   
   //M214
   M2xx_CONVEYOR[11].INPUT_xProtectionRot := A152AP1:3:I.Pt08.Data;
   M2xx_CONVEYOR[11].INPUT_xProtectionFan := xAlwaysON;
   M2xx_CONVEYOR[11].INPUT_xLocalSafetySwitch := A152AP1:10:I.Pt00.Data;
   M2xx_CONVEYOR[11].INPUT_xThermalProbe := A152AP1:10:I.Pt01.Data;
   M2xx_CONVEYOR[11].INPUT_xDriveInhibit := M214_M1_DR.CIPAxisState = 9;
   M2xx_CONVEYOR[11].INPUT_xDriveReady := M214_M1_DR.ServoActionStatus;
   M2xx_CONVEYOR[11].INPUT_xDriveError := M214_M1_DR.AxisFault <> 0 OR M214_M1_DR.ModuleFaults <> 0;
   M2xx_CONVEYOR[11].INPUT_xRotationFeedback := M214_M1_DR.MotionStatus <> 0;
   
   //M215
   M2xx_CONVEYOR[12].INPUT_xProtectionRot := A152AP1:3:I.Pt09.Data;
   M2xx_CONVEYOR[12].INPUT_xProtectionFan := xAlwaysON;
   M2xx_CONVEYOR[12].INPUT_xLocalSafetySwitch := A152AP1:10:I.Pt02.Data;
   M2xx_CONVEYOR[12].INPUT_xThermalProbe := A152AP1:10:I.Pt03.Data;
   M2xx_CONVEYOR[12].INPUT_xDriveInhibit := M215_M1_DR.CIPAxisState = 9;
   M2xx_CONVEYOR[12].INPUT_xDriveReady := M215_M1_DR.ServoActionStatus;
   M2xx_CONVEYOR[12].INPUT_xDriveError := M215_M1_DR.AxisFault <> 0 OR M215_M1_DR.ModuleFaults <> 0;
   M2xx_CONVEYOR[12].INPUT_xRotationFeedback := M215_M1_DR.MotionStatus <> 0;
   
   //M216
   M2xx_CONVEYOR[13].INPUT_xProtectionRot := A152AP1:3:I.Pt10.Data;
   M2xx_CONVEYOR[13].INPUT_xProtectionFan := xAlwaysON;
   M2xx_CONVEYOR[13].INPUT_xLocalSafetySwitch := A152AP1:10:I.Pt04.Data;
   M2xx_CONVEYOR[13].INPUT_xThermalProbe := A152AP1:10:I.Pt05.Data;
   M2xx_CONVEYOR[13].INPUT_xDriveInhibit := M216_M1_DR.CIPAxisState = 9;
   M2xx_CONVEYOR[13].INPUT_xDriveReady := M216_M1_DR.ServoActionStatus;
   M2xx_CONVEYOR[13].INPUT_xDriveError := M216_M1_DR.AxisFault <> 0 OR M216_M1_DR.ModuleFaults <> 0;
   M2xx_CONVEYOR[13].INPUT_xRotationFeedback := M216_M1_DR.MotionStatus <> 0;
   
   //M217
   M2xx_CONVEYOR[14].INPUT_xProtectionRot := A152AP1:3:I.Pt11.Data;
   M2xx_CONVEYOR[14].INPUT_xProtectionFan := xAlwaysON;
   M2xx_CONVEYOR[14].INPUT_xLocalSafetySwitch := A152AP1:10:I.Pt06.Data;
   M2xx_CONVEYOR[14].INPUT_xThermalProbe := A152AP1:10:I.Pt07.Data;
   M2xx_CONVEYOR[14].INPUT_xDriveInhibit := M217_M1_DR.CIPAxisState = 9;
   M2xx_CONVEYOR[14].INPUT_xDriveReady := M217_M1_DR.ServoActionStatus;
   M2xx_CONVEYOR[14].INPUT_xDriveError := M217_M1_DR.AxisFault <> 0 OR M217_M1_DR.ModuleFaults <> 0;
   M2xx_CONVEYOR[14].INPUT_xRotationFeedback := M217_M1_DR.MotionStatus <> 0;
   
   //M218
   M2xx_CONVEYOR[15].INPUT_xProtectionRot := A152AP1:3:I.Pt12.Data;
   M2xx_CONVEYOR[15].INPUT_xProtectionFan := xAlwaysON;
   M2xx_CONVEYOR[15].INPUT_xLocalSafetySwitch := A152AP1:10:I.Pt08.Data;
   M2xx_CONVEYOR[15].INPUT_xThermalProbe := A152AP1:10:I.Pt09.Data;
   M2xx_CONVEYOR[15].INPUT_xDriveInhibit := M218_M1_DR.CIPAxisState = 9;
   M2xx_CONVEYOR[15].INPUT_xDriveReady := M218_M1_DR.ServoActionStatus;
   M2xx_CONVEYOR[15].INPUT_xDriveError := M218_M1_DR.AxisFault <> 0 OR M218_M1_DR.ModuleFaults <> 0;
   M2xx_CONVEYOR[15].INPUT_xRotationFeedback := M218_M1_DR.MotionStatus <> 0;
   
   //M219
   M2xx_CONVEYOR[16].INPUT_xProtectionRot := A152AP1:3:I.Pt13.Data;
   M2xx_CONVEYOR[16].INPUT_xProtectionFan := xAlwaysON;
   M2xx_CONVEYOR[16].INPUT_xLocalSafetySwitch := A152AP1:10:I.Pt10.Data;
   M2xx_CONVEYOR[16].INPUT_xThermalProbe := A152AP1:10:I.Pt11.Data;
   M2xx_CONVEYOR[16].INPUT_xDriveInhibit := M219_M1_DR.CIPAxisState = 9;
   M2xx_CONVEYOR[16].INPUT_xDriveReady := M219_M1_DR.ServoActionStatus;
   M2xx_CONVEYOR[16].INPUT_xDriveError := M219_M1_DR.AxisFault <> 0 OR M219_M1_DR.ModuleFaults <> 0;
   M2xx_CONVEYOR[16].INPUT_xRotationFeedback := M219_M1_DR.MotionStatus <> 0;
   
   //M301M1
   M2xx_CONVEYOR[17].INPUT_xProtectionRot := A152AP1:3:I.Pt14.Data;
   M2xx_CONVEYOR[17].INPUT_xProtectionFan := xAlwaysON;
   M2xx_CONVEYOR[17].INPUT_xLocalSafetySwitch := A152AP1:10:I.Pt12.Data;
   M2xx_CONVEYOR[17].INPUT_xThermalProbe := A152AP1:10:I.Pt13.Data;
   M2xx_CONVEYOR[17].INPUT_xDriveInhibit := M301_M1_DR.CIPAxisState = 9;
   M2xx_CONVEYOR[17].INPUT_xDriveReady := M301_M1_DR.ServoActionStatus;
   M2xx_CONVEYOR[17].INPUT_xDriveError := M301_M1_DR.AxisFault <> 0 OR M301_M1_DR.ModuleFaults <> 0;
   M2xx_CONVEYOR[17].INPUT_xRotationFeedback := M301_M1_DR.MotionStatus <> 0;
   
   
   //M301M2
   M2xx_CONVEYOR[18].INPUT_xProtectionRot := A152AP1:3:I.Pt15.Data;
   M2xx_CONVEYOR[18].INPUT_xProtectionFan := xAlwaysON;
   M2xx_CONVEYOR[18].INPUT_xLocalSafetySwitch := A152AP1:10:I.Pt14.Data;
   M2xx_CONVEYOR[18].INPUT_xThermalProbe := A152AP1:10:I.Pt15.Data;
   M2xx_CONVEYOR[18].INPUT_xDriveInhibit := M301_M2_DR.CIPAxisState = 9;
   M2xx_CONVEYOR[18].INPUT_xDriveReady := M301_M2_DR.ServoActionStatus;
   M2xx_CONVEYOR[18].INPUT_xDriveError := M301_M2_DR.AxisFault <> 0 OR M301_M2_DR.ModuleFaults <> 0;
   M2xx_CONVEYOR[18].INPUT_xRotationFeedback := M301_M2_DR.MotionStatus <> 0;
   
   
   //M220
   M2xx_CONVEYOR[19].INPUT_xProtectionRot := A152AP1:4:I.Pt00.Data;
   M2xx_CONVEYOR[19].INPUT_xProtectionFan := xAlwaysON;
   M2xx_CONVEYOR[19].INPUT_xLocalSafetySwitch := A152AP1:11:I.Pt00.Data;
   M2xx_CONVEYOR[19].INPUT_xThermalProbe := A152AP1:11:I.Pt01.Data;
   M2xx_CONVEYOR[19].INPUT_xDriveInhibit := M220_M1_DR.CIPAxisState = 9;
   M2xx_CONVEYOR[19].INPUT_xDriveReady := M220_M1_DR.ServoActionStatus;
   M2xx_CONVEYOR[19].INPUT_xDriveError := M220_M1_DR.AxisFault <> 0 OR M220_M1_DR.ModuleFaults <> 0;
   M2xx_CONVEYOR[19].INPUT_xRotationFeedback := M220_M1_DR.MotionStatus <> 0;
   
   
   // MAPPING PREVIOUS PROGRAM INPUTS
   
   //ALARM RESET
   I[16].9 := A152AP1:11:I.Pt08.Data;; //VMCC MB Alarm Silence
   I[16].10 := A152AP1:11:I.Pt09.Data;; //VMCC MB Alarm Reset
   
   //ISRA 5D
   I[16].0 := A152AP1:12:I.Pt00.Data; //ISRA 5D 24 VDC OK
   I[16].4 := A152AP1:11:I.Pt06.Data; //ISRA 5D 12 VDC OK
   I[16].5 := A152AP1:11:I.Pt07.Data; //ISRA 5D SYSTEM OK
   I[16].6 := A152AP1:11:I.Pt15.Data; //ISRA 5D System Warning
   I[16].7 := A152AP1:11:I.Pt12.Data; //ISRA 5D System Error 1
   I[16].8 := A152AP1:11:I.Pt13.Data; //ISRA 5D System Error 2
   I[16].14 := A152AP1:11:I.Pt14.Data; //ISRA 5D System Crossbreak
   
   //CHILLED WATER & SUB SURFACE
   I[17].1 := A152AP1:12:I.Pt01.Data; //South Chilled Water Blower Off PB I02105
   I[17].2 := A152AP1:12:I.Pt02.Data; //North Subsurface Cutter Alarm Signal
   I[17].3 := A152AP1:12:I.Pt03.Data; //South Subsurface Cutter Alarm Signal
   I[17].4 := A152AP1:12:I.Pt04.Data; //South Chilled Water Blower On PB I02104
   I[17].5 := A152AP1:12:I.Pt05.Data; //South Chilled Water Blower Off PB I02105
   I[17].7 := A152AP1:12:I.Pt07.Data; //South Chilled Water Blower VFD is Running Without Faults
   I[17].10 := A152AP1:12:I.Pt10.Data; //North Chilled Water Blower On PB I02112
   I[17].11 := A152AP1:12:I.Pt11.Data; //North Chilled Water Blower Off PB I02113
   I[17].13 := A152AP1:12:I.Pt13.Data; //North Chilled Water Blower VFD is Running Without Faults
   
   // CROSSBREAK ZONE 1
   I[24].0 := CB_1CS:0:I.0; //CRSSBRK ZONE 1 North Outside Bypass Switch
   I[24].1 := CB_1CS:0:I.1; //CRSSBRK ZONE 1 North Inside Bypass Switch
   I[24].2 := CB_1CS:0:I.2; //CRSSBRK ZONE 1 South Outside Bypass Switch
   I[24].3 := CB_1CS:0:I.3; //CRSSBRK ZONE 1 South Inside Bypass Switch
   I[24].4 := CB_1CS:0:I.4; //CRSSBRK ZONE 1 North Outside Photo-cell
   I[24].5 := CB_1CS:0:I.5; //CRSSBRK ZONE 1 North Inside Photo-cell
   I[24].6 := CB_1CS:0:I.6; //CRSSBRK ZONE 1 South Outside Photo-cell
   I[24].7 := CB_1CS:0:I.7; //CRSSBRK ZONE 1 South Inside Photo-cell
   I[24].8 := CB_1CS:0:I.8; //Cullet System M37B Fwd Direction Selector (Outside)
   I[24].9 := CB_1CS:0:I.9; //Cullet System M37B Rev Direction Selector (Outside)
   I[24].10 := CB_1CS:0:I.10; //Cullet System M47B Fwd Direction Selector (Outside)
   I[24].11 := CB_1CS:0:I.11; //Cullet System M47B Rev Direction Selector (Outside)
   I[24].12 := CB_1CS:0:I.12; //Diverter Position Selector At Cullet Op Panel (Input from cullet belts 51 running)
   I[24].13 := CB_1CS:0:I.13; //(Input from cullet belts 52 running)
   I[24].14 := CB_1CS:0:I.14; //spare
   I[24].15 := CB_1CS:0:I.15; //spare
   
   // CROSSBREAK ZONE 2
   I[26].0 := CB_2CS:0:I.0; //CRSSBRK ZONE 2 North Outside Bypass Switch
   I[26].1 := CB_2CS:0:I.1; //CRSSBRK ZONE 2 North Inside Bypass Switch
   I[26].2 := CB_2CS:0:I.2; //CRSSBRK ZONE 2 South Outside Bypass Switch
   I[26].3 := CB_2CS:0:I.3; //CRSSBRK ZONE 2 South Inside Bypass Switch
   I[26].4 := CB_2CS:0:I.4; //CRSSBRK ZONE 2 North Outside Photo-cell
   I[26].5 := CB_2CS:0:I.5; //CRSSBRK ZONE 2 North Inside Photo-cell
   I[26].6 := CB_2CS:0:I.6; //CRSSBRK ZONE 2 South Outside Photo-cell
   I[26].7 := CB_2CS:0:I.7; //CRSSBRK ZONE 2 South Inside Photo-cell
   I[26].8 := CB_2CS:0:I.8; //spare
   I[26].9 := CB_2CS:0:I.9; //spare
   I[26].10 := CB_2CS:0:I.10; //spare
   I[26].11 := CB_2CS:0:I.11; //spare
   I[26].12 := CB_2CS:0:I.12; //spare
   I[26].13 := CB_2CS:0:I.13; //Adapter power ON
   I[26].14 := CB_2CS:0:I.14; //Input power ON
   I[26].15 := CB_2CS:0:I.15; //Output power ON
   
   // CROSSBREAK ZONE 3
   I[28].0 := CB_3CS:0:I.0; //CRSSBRK ZONE 3 North Outside Bypass Switch
   I[28].1 := CB_3CS:0:I.1; //CRSSBRK ZONE 3 North Inside Bypass Switch
   I[28].2 := CB_3CS:0:I.2; //CRSSBRK ZONE 3 South Outside Bypass Switch
   I[28].3 := CB_3CS:0:I.3; //CRSSBRK ZONE 3 South Inside Bypass Switch
   I[28].4 := CB_3CS:0:I.4; //CRSSBRK ZONE 3 North Outside Photo-cell
   I[28].5 := CB_3CS:0:I.5; //CRSSBRK ZONE 3 North Inside Photo-cell
   I[28].6 := CB_3CS:0:I.6; //CRSSBRK ZONE 3 South Outside Photo-cell
   I[28].7 := CB_3CS:0:I.7; //CRSSBRK ZONE 3 South Inside Photo-cell
   I[28].8 := CB_3CS:0:I.8; //spare
   I[28].9 := CB_3CS:0:I.9; //spare
   I[28].10 := CB_3CS:0:I.10; //spare
   I[28].11 := CB_3CS:0:I.11; //spare
   I[28].12 := CB_3CS:0:I.12; //spare
   I[28].13 := CB_3CS:0:I.13; //Adapter power ON
   I[28].14 := CB_3CS:0:I.14; //Input power ON
   I[28].15 := CB_3CS:0:I.15; //Output power ON
   
   // CROSSBREAK ZONE 4 (IMAGE AUTO)
   I[30].0 := CB_4CS:0:I.0; //CRSSBRK ZONE 4 North Outside Bypass Switch
   I[30].1 := CB_4CS:0:I.1; //CRSSBRK ZONE 4 North Inside Bypass Switch
   I[30].2 := CB_4CS:0:I.2; //CRSSBRK ZONE 4 South Outside Bypass Switch
   I[30].3 := CB_4CS:0:I.3; //CRSSBRK ZONE 4 South Inside Bypass Switch
   I[30].4 := CB_4CS:0:I.4; //CRSSBRK ZONE 4 North Outside Photo-cell
   I[30].5 := CB_4CS:0:I.5; //CRSSBRK ZONE 4 North Inside Photo-cell
   I[30].6 := CB_4CS:0:I.6; //CRSSBRK ZONE 4 South Outside Photo-cell
   I[30].7 := CB_4CS:0:I.7; //CRSSBRK ZONE 4 South Inside Photo-cell
   I[30].8 := CB_4CS:0:I.8; //IMAGE AUTO Open Graticule Selector Switch (UP)
   I[30].9 := CB_4CS:0:I.9; //IMAGE AUTO Retro Reflector
   I[30].10 := CB_4CS:0:I.10; //spare
   I[30].11 := CB_4CS:0:I.11; //IMAGE AUTO Cover close Acknowledge Push-button (Silence)
   I[30].12 := CB_4CS:0:I.12; //IMAGE AUTO Retro-cover Closed Prox
   I[30].13 := CB_4CS:0:I.13; //Adapter power ON
   I[30].14 := CB_4CS:0:I.14; //IMAGE AUTO Close Graticule Selector Switch (DOWN)
   I[30].15 := CB_4CS:0:I.15; //Output power ON
   
   // CROSSBREAK ZONE 5 (APC)
   I[32].0 := CB_5CS:0:I.0; //CRSSBRK ZONE 5 North Outside Bypass Switch
   I[32].1 := CB_5CS:0:I.1; //CRSSBRK ZONE 5 North Inside Bypass Switch
   I[32].2 := CB_5CS:0:I.2; //CRSSBRK ZONE 5 South Outside Bypass Switch
   I[32].3 := CB_5CS:0:I.3; //CRSSBRK ZONE 5 South Inside Bypass Switch
   I[32].4 := CB_5CS:0:I.4; //CRSSBRK ZONE 5 North Outside Photo-cell
   I[32].5 := CB_5CS:0:I.5; //CRSSBRK ZONE 5 North Inside Photo-cell
   I[32].6 := CB_5CS:0:I.6; //CRSSBRK ZONE 5 South Outside Photo-cell
   I[32].7 := CB_5CS:0:I.7; //CRSSBRK ZONE 5 South Inside Photo-cell
   I[32].8 := CB_5CS:0:I.8; //APC #1 Reset Button After Crossbreak
   I[32].9 := CB_5CS:0:I.9; //APC Spray system OFF (1=OFF) (0=ON)
   I[32].10 := CB_5CS:0:I.10; //APC #2 Reset Button After Crossbreak changed 22Mar2019TC
   I[32].11 := CB_5CS:0:I.11; //APC Spray System Supply Flow Low (From SMC flow meter)
   I[32].12 := CB_5CS:0:I.12; //spare
   I[32].13 := CB_5CS:0:I.13; //Adapter power ON
   I[32].14 := CB_5CS:0:I.14; //Input power ON
   I[32].15 := CB_5CS:0:I.15; //Output power ON
   
   // MANUAL INSPECTION (LOW-E)
   I[34].0 := MI_6CS:0:I.0; //MANUAL INSPCTN Booth Flaw Push-Button
   I[34].1 := MI_6CS:0:I.1; //MANUAL INSPCTN Booth Reject Push-Button
   I[34].2 := MI_6CS:0:I.2; //MANUAL INSPCTN Quality defect switch (Enable/Inhibit)
   I[34].3 := MI_6CS:0:I.3; //LOW-E Inspection Catwalk: Spray Zone 1 Pushbutton
   I[34].4 := MI_6CS:0:I.4; //LOW-E Inspection Catwalk: Spray Zone 2 Pushbutton
   I[34].5 := MI_6CS:0:I.5; //LOW-E Inspection Catwalk: Spray Zone 3 Pushbutton
   I[34].6 := MI_6CS:0:I.6; //LOW-E Inspection Catwalk: Spray Zone 4 Pushbutton
   I[34].7 := MI_6CS:0:I.7; //LOW-E Inspection Catwalk: Spray Zone 5 Pushbutton
   I[34].8 := MI_6CS:0:I.8; //LOW-E Inspection Catwalk: Pulse Entire Ribbon Pushbutton
   I[34].9 := MI_6CS:0:I.9; //spare
   I[34].10 := MI_6CS:0:I.10; //MANUAL INSPCTN MODE MAN
   I[34].11 := MI_6CS:0:I.11; //MANUAL INSPCTN MODE AUTO
   I[34].12 := MI_6CS:0:I.12; //spare
   I[34].13 := MI_6CS:0:I.13; //Adapter power ON
   I[34].14 := MI_6CS:0:I.14; //Input power ON
   I[34].15 := MI_6CS:0:I.15; //Output power ON
   
   //I[34].10 := A152AP1:11:I.Pt10.Data; // MANUAL INSPECTION MODE MAN
   //I[34].11 := A152AP1:11:I.Pt11.Data; // MANUAL INSPECTION MODE AUTO
   
   //VMCC M1
   I[64].0 := Z200.INPUT_x24VdcVoltageON AND Z200.INPUT_xMainSwitch; //VMCC M1 Drive Contactor Energized
   I[64].1 := Z200.INPUT_xPowerSupply24VLogic1 AND  Z200.INPUT_xPowerSupply24VLogic2; //VMCC1 M1 DC Input Power ON (NOT USED)
   I[64].2 := Z200.INPUT_xPowerSupply24VLogic3 AND  Z200.INPUT_xPowerSupply24VLogic4; //VMCC1 M1 DC Output Power ON (NOT USED)
   //
   I[64].4 := Z200.INPUT_xPowerSupplyOK; //VMCC M1 E-Stop Power ON (NOT USED)
   I[64].5 := Z200.INPUT_xPowerSupplyOK; //VMCC M1 DC Power Supply #1 ON (NOT USED)
   I[64].6 := Z200.INPUT_xPowerSupplyOK; //VMCC M1 DC Power Supply #2 ON (NOT USED)
   //
   I[64].8 := Z200.INPUT_xAlarmSilence; //VMCC M1 Alarm Silence
   I[64].9 := Z200.INPUT_xAlarmReset;	//VMCC M1 Alarm Reset
   I[64].10 := Z200.INPUT_xMainEmergencyON; //VMCC M1 E-Stop Circuit Energized
   I[64].11 := M203DROP.INPUT_xDownPosition; //VMCC M1 Crusher Bar Lowered
   I[64].12 := M203DROP.INPUT_xUpPosition; //VMCC M1 Crusher Bar Raised
   I[64].13 := M203DROP.ST_xOutputEnable; //VMCC M1 Crusher #1 in auto
   I[64].14 := (M203DROP.INPUT_xUpDownPushbuttonOpSide OR M203DROP.INPUT_xUpDownPushbuttonFarSide) AND M203DROP.INPUT_xDownPosition; //VMCC M1 Crusher #1 Manual raise
   I[64].15 := (M203DROP.INPUT_xUpDownPushbuttonOpSide OR M203DROP.INPUT_xUpDownPushbuttonFarSide) AND M203DROP.INPUT_xUpPosition; //VMCC M1 Crusher #1 Manual lower
   
   //VMCC W1 (WASHER)
   I[43].0 := A80AZ1:I.Faulted; //VMCC W1 Upper Brush #1 Drive fault
   I[43].1 := A80AZ1:I.Faulted; //VMCC W1 Lower Brush #1 Drive fault
   I[43].2 := A81AZ1:I.Faulted; //VMCC W1 Upper Brush #2 Drive fault
   I[43].3 := A81AZ1:I.Faulted; //VMCC W1 Lower Brush #2 Drive fault
   
   //PANEL W2 (WASHER)
   I[56].0 := PANEL_W2:0:I.0; //PANEL W2 BRUSH #1 AUTO Sw. Pos.
   I[56].1 := PANEL_W2:0:I.1; //PANEL W2 BRUSH #1 MANUAL Sw. Pos.
   I[56].2 := PANEL_W2:0:I.2; //PANEL W2 BRUSH #1 ON Sw. Pos.
   I[56].3 := PANEL_W2:0:I.3; //PANEL W2 BRUSH #1 OFF Sw. Pos.
   I[56].4 := PANEL_W2:0:I.4; //PANEL W2 BRUSH #2 AUTO Sw. Pos. (NOT USED ANYMORE)
   I[56].5 := PANEL_W2:0:I.5; //PANEL W2 BRUSH #2 MANUAL Sw. Pos. (NOT USED ANYMORE)
   I[56].6 := PANEL_W2:0:I.6; //PANEL W2 BRUSH #2 ON Sw. Pos. (NOT USED ANYMORE)
   I[56].7 := PANEL_W2:0:I.7; //PANEL W2 BRUSH #2 OFF Sw. Pos. (NOT USED ANYMORE)
   I[56].8 := PANEL_W2:0:I.8; //PANEL W2 SPONGE UNIT AUTO Sw. Pos.
   I[56].9 := PANEL_W2:0:I.9; //PANEL W2 SPONGE UNIT MANUAL Sw. Pos.
   I[56].10 := PANEL_W2:0:I.10; //PANEL W2 SPONGE UNIT ON Sw. Pos.
   I[56].11 := PANEL_W2:0:I.11; //PANEL W2 SPONGE UNIT OFF Sw. Pos.
   I[56].12 := PANEL_W2:0:I.12; //PANEL W2 AIR KNIFE AUTO Sw. Pos.
   I[56].13 := PANEL_W2:0:I.13; //PANEL W2 AIR KNIFE MANUAL Sw. Pos.
   I[56].14 := PANEL_W2:0:I.14; //SPARE
   I[56].15 := PANEL_W2:0:I.15; //SPARE
   I[57].0 := PANEL_W2:1:I.0; //PANEL W2 BRUSH #1 UPPER BRUSH CONVERGE Sw. Pos.
   I[57].1 := PANEL_W2:1:I.1; //PANEL W2 BRUSH #1 UPPER BRUSH RETRACT Sw. Pos.
   I[57].2 := PANEL_W2:1:I.2; //PANEL W2 BRUSH #2 UPPER BRUSH CONVERGE Sw. Pos. (NOT USED ANYMORE)
   I[57].3 := PANEL_W2:1:I.3; //PANEL W2 BRUSH #2 UPPER BRUSH RETRACT Sw. Pos. (NOT USED ANYMORE)
   I[57].4 := PANEL_W2:1:I.4; //PANEL W2 SPONGE UNIT UPPER SPONGE CONVERGE Sw. Pos.
   I[57].5 := PANEL_W2:1:I.5; //PANEL W2 SPONGE UNIT UPPER SPONGE RETRACT Sw. Pos.
   I[57].6 := PANEL_W2:1:I.6; //PANEL W2 BRUSH #1 LOWER BRUSH CONVERGE Sw. Pos.
   I[57].7 := PANEL_W2:1:I.7; //PANEL W2 BRUSH #1 LOWER BRUSH RETRACT Sw. Pos.
   I[57].8 := PANEL_W2:1:I.8; //PANEL W2 BRUSH #2 LOWER BRUSH CONVERGE Sw. Pos. (NOT USED ANYMORE)
   I[57].9 := PANEL_W2:1:I.9; //PANEL W2 BRUSH #2 LOWER BRUSH RETRACT Sw. Pos. (NOT USED ANYMORE)
   I[57].10 := PANEL_W2:1:I.10; //PANEL W2 SPONGE UNIT LOWER SPONGE CONVERGE Sw. Pos.
   I[57].11 := PANEL_W2:1:I.11; //PANEL W2 SPONGE UNIT LOWER SPONGE RETRACT Sw. Pos.
   I[57].12 := PANEL_W2:1:I.12; //PANEL W2 AIR KNIFE UNIT #1 CONVERGE Sw. Pos.
   I[57].13 := PANEL_W2:1:I.13; //PANEL W2 AIR KNIFE UNIT #1 RETRACT Sw. Pos.
   I[57].14 := PANEL_W2:1:I.14; //PANEL W2 AIR KNIFE UNIT #2 CONVERGE Sw. Pos.
   I[57].15 := PANEL_W2:1:I.15; //PANEL W2 AIR KNIFE UNIT #2 RETRACT Sw. Pos.
   I[58].0 := PANEL_W2:2:I.0; //PANEL W2 Cross break Reset Push-button
   I[58].1 := PANEL_W2:2:I.1; //PANEL W2 WATER SPRAYERS AUTO  Sw. Pos.
   I[58].2 := PANEL_W2:2:I.2; //PANEL W2 WATER SPRAYERS MANUAL  Sw. Pos.
   I[58].3 := PANEL_W2:2:I.3; //PANEL W2 WATER SPRAYERS ON  Sw. Pos.
   I[58].4 := PANEL_W2:2:I.4; //PANEL W2 WATER SPRAYERS OFF  Sw. Pos.
   I[58].5 := PANEL_W2:2:I.5; //PANEL W2 SELECTOR SWITCH CITRIC ACID WASHER ON (# W2) (NOT USED ANYMORE)
   I[58].6 := PANEL_W2:2:I.6; //PANEL W2 SELECTOR SWITCH CITRIC ACID WASHER OFF (# W2) (NOT USED ANYMORE)
   I[58].7 := PANEL_W2:2:I.7; //PANEL W2 AIR KNIFE BLOWER MODE ON SS PANEL #W2
   I[58].8 := PANEL_W2:2:I.8; //PANEL W2 AIR KNIFE BLOWER MODE OFF SS PANEL #W2
   I[58].9 := PANEL_W2:2:I.9; //SPARE
   I[58].10 := PANEL_W2:2:I.10; //SPARE
   I[58].11 := PANEL_W2:2:I.11; //SPARE
   I[58].12 := PANEL_W2:2:I.12; //SPARE
   I[58].13 := PANEL_W2:2:I.13; //SPARE
   I[58].14 := PANEL_W2:2:I.14; //SPARE
   I[58].15 := PANEL_W2:2:I.15; //SPARE
   
   //PANEL W3 (WASHER)
   I[60].0 := PANEL_W3:0:I.0; //PANEL W3 BRUSH #1 AUTO Sw. Pos.
   I[60].1 := PANEL_W3:0:I.1; //PANEL W3 BRUSH #1 MANUAL Sw. Pos.
   I[60].2 := PANEL_W3:0:I.2; //PANEL W3 BRUSH #1 ON Sw. Pos.
   I[60].3 := PANEL_W3:0:I.3; //PANEL W3 BRUSH #1 OFF Sw. Pos.
   I[60].4 := PANEL_W3:0:I.4; //PANEL W3 BRUSH #2 AUTO Sw. Pos. (NOT USED ANYMORE)
   I[60].5 := PANEL_W3:0:I.5; //PANEL W3 BRUSH #2 MANUAL Sw. Pos. (NOT USED ANYMORE)
   I[60].6 := PANEL_W3:0:I.6; //PANEL W3 BRUSH #2 ON Sw. Pos. (NOT USED ANYMORE)
   I[60].7 := PANEL_W3:0:I.7; //PANEL W3 BRUSH #2 OFF Sw. Pos. (NOT USED ANYMORE)
   I[60].8 := PANEL_W3:0:I.8; //PANEL W3 SPONGE UNIT AUTO Sw. Pos.
   I[60].9 := PANEL_W3:0:I.9; //PANEL W3 SPONGE UNIT MANUAL Sw. Pos.
   I[60].10 := PANEL_W3:0:I.10; //PANEL W3 SPONGE UNIT ON Sw. Pos.
   I[60].11 := PANEL_W3:0:I.11; //PANEL W3 SPONGE UNIT OFF Sw. Pos.
   I[60].12 := PANEL_W3:0:I.12; //PANEL W3 AIR KNIFE AUTO Sw. Pos.
   I[60].13 := PANEL_W3:0:I.13; //PANEL W3 AIR KNIFE MANUAL Sw. Pos.
   I[60].14 := PANEL_W3:0:I.14; //PANEL W3 JOG SPONGE ROLL FORWARD
   I[60].15 := PANEL_W3:0:I.15; //SPARE
   I[61].0 := PANEL_W3:1:I.0; //PANEL W3 BRUSH #1 UPPER BRUSH CONVERGE Sw. Pos.
   I[61].1 := PANEL_W3:1:I.1; //PANEL W3 BRUSH #1 UPPER BRUSH RETRACT Sw. Pos.
   I[61].2 := PANEL_W3:1:I.2; //PANEL W3 BRUSH #2 UPPER BRUSH CONVERGE Sw. Pos. (NOT USED ANYMORE)
   I[61].3 := PANEL_W3:1:I.3; //PANEL W3 BRUSH #2 UPPER BRUSH RETRACT Sw. Pos. (NOT USED ANYMORE)
   I[61].4 := PANEL_W3:1:I.4; //PANEL W3 SPONGE UNIT UPPER SPONGE CONVERGE Sw. Pos.
   I[61].5 := PANEL_W3:1:I.5; //PANEL W3 SPONGE UNIT UPPER SPONGE RETRACT Sw. Pos.
   I[61].6 := PANEL_W3:1:I.6; //PANEL W3 BRUSH #1 LOWER BRUSH CONVERGE Sw. Pos.
   I[61].7 := PANEL_W3:1:I.7; //PANEL W3 BRUSH #1 LOWER BRUSH RETRACT Sw. Pos.
   I[61].8 := PANEL_W3:1:I.8; //PANEL W3 BRUSH #2 LOWER BRUSH CONVERGE Sw. Pos. (NOT USED ANYMORE)
   I[61].9 := PANEL_W3:1:I.9; //PANEL W3 BRUSH #2 LOWER BRUSH RETRACT Sw. Pos. (NOT USED ANYMORE)
   I[61].10 := PANEL_W3:1:I.10; //PANEL W3 SPONGE UNIT LOWER SPONGE CONVERGE Sw. Pos.
   I[61].11 := PANEL_W3:1:I.11; //PANEL W3 SPONGE UNIT LOWER SPONGE RETRACT Sw. Pos.
   I[61].12 := PANEL_W3:1:I.12; //PANEL W3 AIR KNIFE UNIT #1 CONVERGE Sw. Pos.
   I[61].13 := PANEL_W3:1:I.13; //PANEL W3 AIR KNIFE UNIT #1 RETRACT Sw. Pos.
   I[61].14 := PANEL_W3:1:I.14; //PANEL W3 AIR KNIFE UNIT #2 CONVERGE Sw. Pos.
   I[61].15 := PANEL_W3:1:I.15; //PANEL W3 AIR KNIFE UNIT #2 RETRACT Sw. Pos.
   I[62].0 := PANEL_W3:1:I.0; //PANEL W3 Cross break Reset Push-button
   I[62].1 := PANEL_W3:2:I.1; //PANEL W3 WATER SPRAYERS AUTO  Sw. Pos.
   I[62].2 := PANEL_W3:2:I.2; //PANEL W3 WATER SPRAYERS MANUAL  Sw. Pos.
   I[62].3 := PANEL_W3:2:I.3; //PANEL W3 WATER SPRAYERS ON  Sw. Pos.
   I[62].4 := PANEL_W3:2:I.4; //PANEL W3 WATER SPRAYERS OFF  Sw. Pos.
   I[62].5 := PANEL_W3:2:I.5; //PANEL W3 SELECTOR SWITCH CITRIC ACID WASHER ON (# W3) (NOT USED ANYMORE)
   I[62].6 := PANEL_W3:2:I.6; //PANEL W3 SELECTOR SWITCH CITRIC ACID WASHER OFF (# W3) (NOT USED ANYMORE)
   I[62].7 := PANEL_W3:2:I.7; //PANEL W3 AIR KNIFE BLOWER MODE ON SS PANEL #W3
   I[62].8 := PANEL_W3:2:I.8; //PANEL W3 AIR KNIFE BLOWER MODE OFF SS PANEL #W3
   I[62].9 := PANEL_W3:2:I.9; //SPARE
   I[62].10 := PANEL_W3:2:I.10; //SPARE
   I[62].11 := PANEL_W3:2:I.11; //SPARE
   I[62].12 := PANEL_W3:2:I.12; //SPARE
   I[62].13 := PANEL_W3:2:I.13; //SPARE
   I[62].14 := PANEL_W3:2:I.14; //SPARE
   I[62].15 := PANEL_W3:2:I.15; //SPARE
   
   
   //CONSUMED
   
   I[112] := From_Cullet[0];
   I[113] := From_Cullet[1];
   I[114] := From_Cullet[2];
   I[115] := From_Cullet[3];
   I[116] := From_Cullet[4];
   I[117] := From_Cullet[5];
   I[118] := From_Cullet[6];
   I[119] := From_Cullet[7];
   
   /*
   
   I[112] := ConsumedFromCullet.iCULLETtoMB_1;
   I[113] := ConsumedFromCullet.iCULLETtoMB_2;
   I[114] := ConsumedFromCullet.iCULLETtoMB_3;
   I[115] := ConsumedFromCullet.iCULLETtoMB_4;
   I[116] := ConsumedFromCullet.iCULLETtoMB_5;
   I[117] := ConsumedFromCullet.iCULLETtoMB_6;
   I[118] := ConsumedFromCullet.iCULLETtoMB_7;
   I[119] := ConsumedFromCullet.iCULLETtoMB_8;
   
   */
   
   I[120] := ConsumedFromMCC1300.iM2toMB_1;
   I[121] := ConsumedFromMCC1300.iM2toMB_2;
   I[122] := ConsumedFromMCC1300.iM2toMB_3;
   I[123] := ConsumedFromMCC1300.iM2toMB_4;
   I[124] := ConsumedFromMCC1300.iM2toMB_5;
   I[125] := ConsumedFromMCC1300.iM2toMB_6;
   I[126] := ConsumedFromMCC1300.iM2toMB_7;
   I[127] := ConsumedFromMCC1300.iM2toMB_8;
   
   
   //DRIVE
   
   
   //MOTION
   
   COP(M301_M1_DR_OUT_MAJ,M301_M1_DR_IN_MAJ,1);
   M301_M1_DR_IN_MAR.EN := M301_M1_DR_OUT_MAR.EN;
   M301_M1_DR_IN_MAR.PC := M301_M1_DR_OUT_MAR.PC;
   COP(M301_M1_DR_OUT_MAM,M301_M1_DR_IN_MAM,1);
   COP(M301_M1_DR_OUT_MAS,M301_M1_DR_IN_MAS,1);
   COP(M301_M1_DR_OUT_MRP,M301_M1_DR_IN_MRP,1);
   COP(M301_M1_DR_OUT_MCD,M301_M1_DR_IN_MCD,1);
   
   COP(M301_M2_DR_OUT_MAJ,M301_M2_DR_IN_MAJ,1);
   M301_M2_DR_IN_MAR.EN := M301_M2_DR_OUT_MAR.EN;
   M301_M2_DR_IN_MAR.PC := M301_M2_DR_OUT_MAR.PC;
   COP(M301_M2_DR_OUT_MAM,M301_M2_DR_IN_MAM,1);
   COP(M301_M2_DR_OUT_MAS,M301_M2_DR_IN_MAS,1);
   COP(M301_M2_DR_OUT_MRP,M301_M2_DR_IN_MRP,1);
   COP(M301_M2_DR_OUT_MCD,M301_M2_DR_IN_MCD,1);
   
   COP(M202_M1_DR_OUT_MAJ,M202_M1_DR_IN_MAJ,1);
   M202_M1_DR_IN_MAR.EN := M202_M1_DR_OUT_MAR.EN;
   M202_M1_DR_IN_MAR.PC := M202_M1_DR_OUT_MAR.PC;
   COP(M202_M1_DR_OUT_MAM,M202_M1_DR_IN_MAM,1);
   COP(M202_M1_DR_OUT_MAS,M202_M1_DR_IN_MAS,1);
   COP(M202_M1_DR_OUT_MRP,M202_M1_DR_IN_MRP,1);
   COP(M202_M1_DR_OUT_MCD,M202_M1_DR_IN_MCD,1);
   
   COP(M203_M1_DR_OUT_MAJ,M203_M1_DR_IN_MAJ,1);
   M203_M1_DR_IN_MAR.EN := M203_M1_DR_OUT_MAR.EN;
   M203_M1_DR_IN_MAR.PC := M203_M1_DR_OUT_MAR.PC;
   COP(M203_M1_DR_OUT_MAM,M203_M1_DR_IN_MAM,1);
   COP(M203_M1_DR_OUT_MAS,M203_M1_DR_IN_MAS,1);
   COP(M203_M1_DR_OUT_MRP,M203_M1_DR_IN_MRP,1);
   COP(M203_M1_DR_OUT_MCD,M203_M1_DR_IN_MCD,1);
   
   COP(M204_M1_DR_OUT_MAJ,M204_M1_DR_IN_MAJ,1);
   M204_M1_DR_IN_MAR.EN := M204_M1_DR_OUT_MAR.EN;
   M204_M1_DR_IN_MAR.PC := M204_M1_DR_OUT_MAR.PC;
   COP(M204_M1_DR_OUT_MAM,M204_M1_DR_IN_MAM,1);
   COP(M204_M1_DR_OUT_MAS,M204_M1_DR_IN_MAS,1);
   COP(M204_M1_DR_OUT_MRP,M204_M1_DR_IN_MRP,1);
   COP(M204_M1_DR_OUT_MCD,M204_M1_DR_IN_MCD,1);
   
   COP(M206_M1_DR_OUT_MAJ,M206_M1_DR_IN_MAJ,1);
   M206_M1_DR_IN_MAR.EN := M206_M1_DR_OUT_MAR.EN;
   M206_M1_DR_IN_MAR.PC := M206_M1_DR_OUT_MAR.PC;
   COP(M206_M1_DR_OUT_MAM,M206_M1_DR_IN_MAM,1);
   COP(M206_M1_DR_OUT_MAS,M206_M1_DR_IN_MAS,1);
   COP(M206_M1_DR_OUT_MRP,M206_M1_DR_IN_MRP,1);
   COP(M206_M1_DR_OUT_MCD,M206_M1_DR_IN_MCD,1);
   
   COP(M207_M1_DR_OUT_MAJ,M207_M1_DR_IN_MAJ,1);
   M207_M1_DR_IN_MAR.EN := M207_M1_DR_OUT_MAR.EN;
   M207_M1_DR_IN_MAR.PC := M207_M1_DR_OUT_MAR.PC;
   COP(M207_M1_DR_OUT_MAM,M207_M1_DR_IN_MAM,1);
   COP(M207_M1_DR_OUT_MAS,M207_M1_DR_IN_MAS,1);
   COP(M207_M1_DR_OUT_MRP,M207_M1_DR_IN_MRP,1);
   COP(M207_M1_DR_OUT_MCD,M207_M1_DR_IN_MCD,1);
   
   COP(M208_M1_DR_OUT_MAJ,M208_M1_DR_IN_MAJ,1);
   M208_M1_DR_IN_MAR.EN := M208_M1_DR_OUT_MAR.EN;
   M208_M1_DR_IN_MAR.PC := M208_M1_DR_OUT_MAR.PC;
   COP(M208_M1_DR_OUT_MAM,M208_M1_DR_IN_MAM,1);
   COP(M208_M1_DR_OUT_MAS,M208_M1_DR_IN_MAS,1);
   COP(M208_M1_DR_OUT_MRP,M208_M1_DR_IN_MRP,1);
   COP(M208_M1_DR_OUT_MCD,M208_M1_DR_IN_MCD,1);
   
   COP(M209_M1_DR_OUT_MAJ,M209_M1_DR_IN_MAJ,1);
   M209_M1_DR_IN_MAR.EN := M209_M1_DR_OUT_MAR.EN;
   M209_M1_DR_IN_MAR.PC := M209_M1_DR_OUT_MAR.PC;
   COP(M209_M1_DR_OUT_MAM,M209_M1_DR_IN_MAM,1);
   COP(M209_M1_DR_OUT_MAS,M209_M1_DR_IN_MAS,1);
   COP(M209_M1_DR_OUT_MRP,M209_M1_DR_IN_MRP,1);
   COP(M209_M1_DR_OUT_MCD,M209_M1_DR_IN_MCD,1);
   
   COP(M210_M1_DR_OUT_MAJ,M210_M1_DR_IN_MAJ,1);
   M210_M1_DR_IN_MAR.EN := M210_M1_DR_OUT_MAR.EN;
   M210_M1_DR_IN_MAR.PC := M210_M1_DR_OUT_MAR.PC;
   COP(M210_M1_DR_OUT_MAM,M210_M1_DR_IN_MAM,1);
   COP(M210_M1_DR_OUT_MAS,M210_M1_DR_IN_MAS,1);
   COP(M210_M1_DR_OUT_MRP,M210_M1_DR_IN_MRP,1);
   COP(M210_M1_DR_OUT_MCD,M210_M1_DR_IN_MCD,1);
   
   COP(M211_M1_DR_OUT_MAJ,M211_M1_DR_IN_MAJ,1);
   M211_M1_DR_IN_MAR.EN := M211_M1_DR_OUT_MAR.EN;
   M211_M1_DR_IN_MAR.PC := M211_M1_DR_OUT_MAR.PC;
   COP(M211_M1_DR_OUT_MAM,M211_M1_DR_IN_MAM,1);
   COP(M211_M1_DR_OUT_MAS,M211_M1_DR_IN_MAS,1);
   COP(M211_M1_DR_OUT_MRP,M211_M1_DR_IN_MRP,1);
   COP(M211_M1_DR_OUT_MCD,M211_M1_DR_IN_MCD,1);
   
   COP(M212_M1_DR_OUT_MAJ,M212_M1_DR_IN_MAJ,1);
   M212_M1_DR_IN_MAR.EN := M212_M1_DR_OUT_MAR.EN;
   M212_M1_DR_IN_MAR.PC := M212_M1_DR_OUT_MAR.PC;
   COP(M212_M1_DR_OUT_MAM,M212_M1_DR_IN_MAM,1);
   COP(M212_M1_DR_OUT_MAS,M212_M1_DR_IN_MAS,1);
   COP(M212_M1_DR_OUT_MRP,M212_M1_DR_IN_MRP,1);
   COP(M212_M1_DR_OUT_MCD,M212_M1_DR_IN_MCD,1);
   
   COP(M213_M1_DR_OUT_MAJ,M213_M1_DR_IN_MAJ,1);
   M213_M1_DR_IN_MAR.EN := M213_M1_DR_OUT_MAR.EN;
   M213_M1_DR_IN_MAR.PC := M213_M1_DR_OUT_MAR.PC;
   COP(M213_M1_DR_OUT_MAM,M213_M1_DR_IN_MAM,1);
   COP(M213_M1_DR_OUT_MAS,M213_M1_DR_IN_MAS,1);
   COP(M213_M1_DR_OUT_MRP,M213_M1_DR_IN_MRP,1);
   COP(M213_M1_DR_OUT_MCD,M213_M1_DR_IN_MCD,1);
   
   COP(M213A_M1_DR_OUT_MAJ,M213A_M1_DR_IN_MAJ,1);
   M213A_M1_DR_IN_MAR.EN := M213A_M1_DR_OUT_MAR.EN;
   M213A_M1_DR_IN_MAR.PC := M213A_M1_DR_OUT_MAR.PC;
   COP(M213A_M1_DR_OUT_MAM,M213A_M1_DR_IN_MAM,1);
   COP(M213A_M1_DR_OUT_MAS,M213A_M1_DR_IN_MAS,1);
   COP(M213A_M1_DR_OUT_MRP,M213A_M1_DR_IN_MRP,1);
   COP(M213A_M1_DR_OUT_MCD,M213A_M1_DR_IN_MCD,1);
   
   COP(M213B_M1_DR_OUT_MAJ,M213B_M1_DR_IN_MAJ,1);
   M213B_M1_DR_IN_MAR.EN := M213B_M1_DR_OUT_MAR.EN;
   M213B_M1_DR_IN_MAR.PC := M213B_M1_DR_OUT_MAR.PC;
   COP(M213B_M1_DR_OUT_MAM,M213B_M1_DR_IN_MAM,1);
   COP(M213B_M1_DR_OUT_MAS,M213B_M1_DR_IN_MAS,1);
   COP(M213B_M1_DR_OUT_MRP,M213B_M1_DR_IN_MRP,1);
   COP(M213B_M1_DR_OUT_MCD,M213B_M1_DR_IN_MCD,1);
   
   COP(M214_M1_DR_OUT_MAJ,M214_M1_DR_IN_MAJ,1);
   M214_M1_DR_IN_MAR.EN := M214_M1_DR_OUT_MAR.EN;
   M214_M1_DR_IN_MAR.PC := M214_M1_DR_OUT_MAR.PC;
   COP(M214_M1_DR_OUT_MAM,M214_M1_DR_IN_MAM,1);
   COP(M214_M1_DR_OUT_MAS,M214_M1_DR_IN_MAS,1);
   COP(M214_M1_DR_OUT_MRP,M214_M1_DR_IN_MRP,1);
   COP(M214_M1_DR_OUT_MCD,M214_M1_DR_IN_MCD,1);